REGION Network 189: CARRIER SPACING FAULT
   RUNG wire#powerrail
      Contact( "reset" )
      Contact( "EMS".Carrier[5].SDC_OUT.Faults.CarrierSpacingFault )
      wire#w1
      Coil( "DB302_HMI_Faults".Carrier5_Faults_2.%X2 )
   END_RUNG
   RUNG wire#powerrail
      Contact( "DB302_HMI_Faults".Carrier5_Faults_2.%X2 )
      I_Contact( "EMS_Fault_Reset" )
   END_RUNG wire#w1
   // the same network as SCL:
   "DB302_HMI_Faults".Carrier5_Faults_2.%X2 := ("reset" AND "EMS".Carrier[5].SDC_OUT.Faults.CarrierSpacingFault) OR ("DB302_HMI_Faults".Carrier5_Faults_2.%X2 AND NOT "EMS_Fault_Reset");
END_REGION

REGION Network 190: DUPLICATE CARRIER NUMBER FAULT
   RUNG wire#powerrail
      Contact( "reset" )
      Contact( "EMS".Carrier[5].SDC_OUT.Faults.DuplicateCarrierFault )
      wire#w1
      Coil( "DB302_HMI_Faults".Carrier5_Faults_2.%X3 )
   END_RUNG
   RUNG wire#powerrail
      Contact( "DB302_HMI_Faults".Carrier5_Faults_2.%X3 )
      I_Contact( "EMS_Fault_Reset" )
   END_RUNG wire#w1
   // the same network as SCL:
   "DB302_HMI_Faults".Carrier5_Faults_2.%X3 := ("reset" AND "EMS".Carrier[5].SDC_OUT.Faults.DuplicateCarrierFault) OR ("DB302_HMI_Faults".Carrier5_Faults_2.%X3 AND NOT "EMS_Fault_Reset");
END_REGION

REGION Network 191: PRODUCTION HOLD PB NOT RESET
   RUNG wire#powerrail
      Contact( "reset" )
      { S7_Templates := "SrcType := Word" } EQ_Contact(in1 := "DB101_DB_SDC_FAULTS".Carrier_Fault[5], in2 := 103)
      Coil( "DB302_HMI_Faults".Carrier5_Faults_3.%X14 )
   END_RUNG
   // the same network as SCL:
   "DB302_HMI_Faults".Carrier5_Faults_3.%X14 := "reset" AND ("DB101_DB_SDC_FAULTS".Carrier_Fault[5] = 103);
END_REGION

REGION Network 192: CARRIER FAULTS MASKED
   Label( C05_Comm_Flt )
   RUNG wire#powerrail
      Contact( "EMS".Carrier[5].FaultsMasked )
      Coil( "DB302_HMI_Faults".Carrier5_Faults_3.%X15 )
   END_RUNG
   // the same network as SCL:
   C05_Comm_Flt:
   "DB302_HMI_Faults".Carrier5_Faults_3.%X15 := "EMS".Carrier[5].FaultsMasked;
END_REGION

REGION Network 193: CARRIER 6 FAULTS
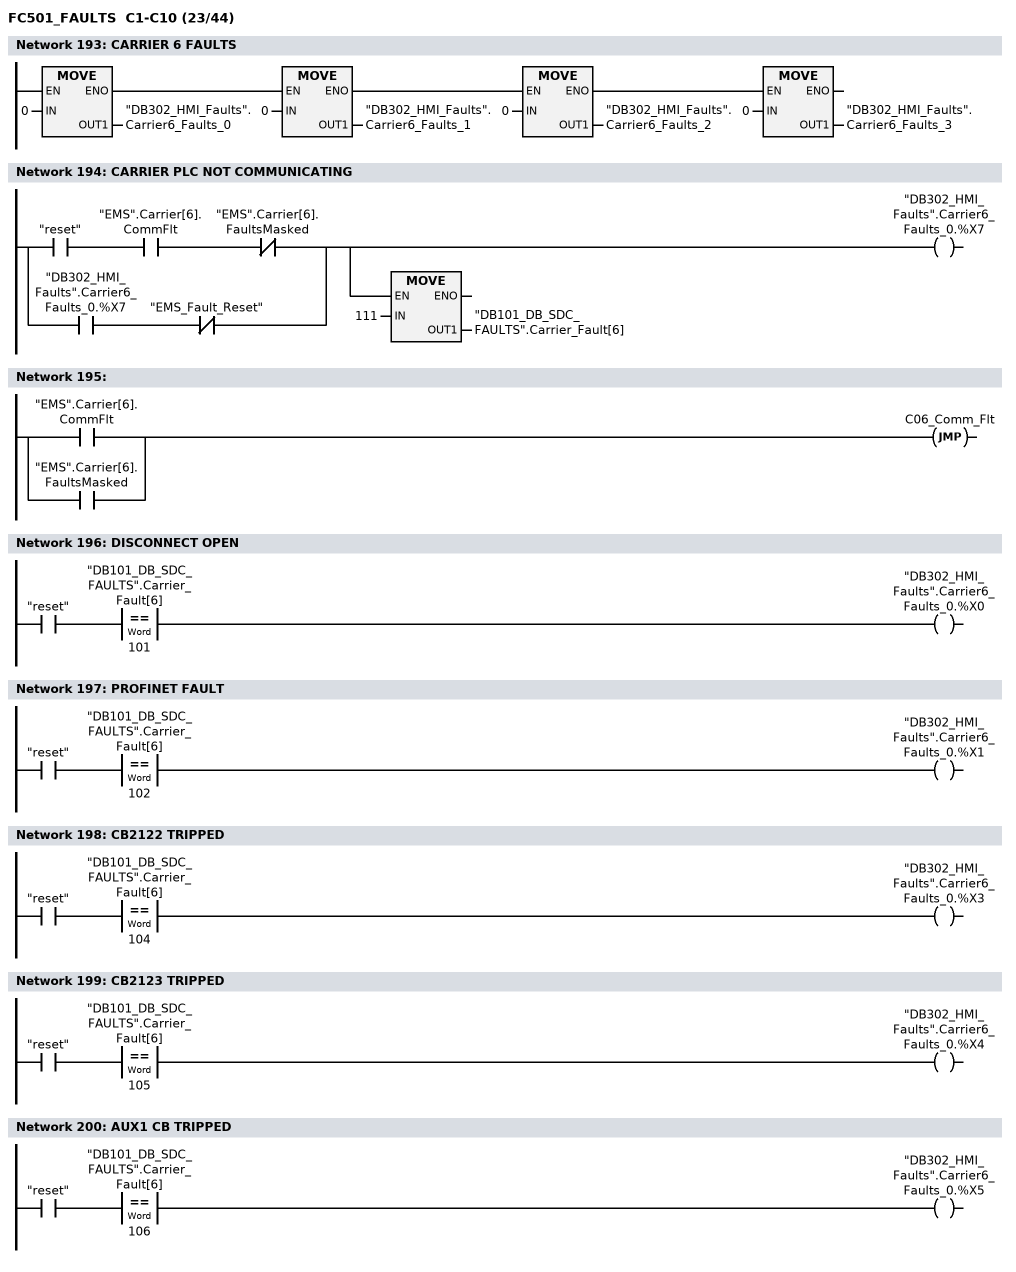
   RUNG wire#powerrail
      Move(in := 0, out1 => "DB302_HMI_Faults".Carrier6_Faults_0)
      Move(in := 0, out1 => "DB302_HMI_Faults".Carrier6_Faults_1)
      Move(in := 0, out1 => "DB302_HMI_Faults".Carrier6_Faults_2)
      Move(in := 0, out1 => "DB302_HMI_Faults".Carrier6_Faults_3)
   END_RUNG
   // the same network as SCL:
   "DB302_HMI_Faults".Carrier6_Faults_0 := 0;
   "DB302_HMI_Faults".Carrier6_Faults_1 := 0;
   "DB302_HMI_Faults".Carrier6_Faults_2 := 0;
   "DB302_HMI_Faults".Carrier6_Faults_3 := 0;
END_REGION

REGION Network 194: CARRIER PLC NOT COMMUNICATING
   RUNG wire#powerrail
      Contact( "reset" )
      Contact( "EMS".Carrier[6].CommFlt )
      I_Contact( "EMS".Carrier[6].FaultsMasked )
      wire#w1
      Coil( "DB302_HMI_Faults".Carrier6_Faults_0.%X7 )
   END_RUNG
   RUNG wire#powerrail
      Contact( "DB302_HMI_Faults".Carrier6_Faults_0.%X7 )
      I_Contact( "EMS_Fault_Reset" )
   END_RUNG wire#w1
   RUNG wire#w1
      Move(in := 111, out1 => "DB101_DB_SDC_FAULTS".Carrier_Fault[6])
   END_RUNG
   // the same network as SCL:
   "DB302_HMI_Faults".Carrier6_Faults_0.%X7 := ("reset" AND "EMS".Carrier[6].CommFlt AND NOT "EMS".Carrier[6].FaultsMasked) OR ("DB302_HMI_Faults".Carrier6_Faults_0.%X7 AND NOT "EMS_Fault_Reset");
   IF "DB302_HMI_Faults".Carrier6_Faults_0.%X7 THEN "DB101_DB_SDC_FAULTS".Carrier_Fault[6] := 111; END_IF;
END_REGION

REGION Network 195
   RUNG wire#powerrail
      Contact( "EMS".Carrier[6].CommFlt )
      wire#w1
      JumpCoil( C06_Comm_Flt )
   END_RUNG
   RUNG wire#powerrail
      Contact( "EMS".Carrier[6].FaultsMasked )
   END_RUNG wire#w1
   // the same network as SCL:
   IF "EMS".Carrier[6].CommFlt OR "EMS".Carrier[6].FaultsMasked THEN GOTO C06_Comm_Flt; END_IF;
END_REGION

REGION Network 196: DISCONNECT OPEN
   RUNG wire#powerrail
      Contact( "reset" )
      { S7_Templates := "SrcType := Word" } EQ_Contact(in1 := "DB101_DB_SDC_FAULTS".Carrier_Fault[6], in2 := 101)
      Coil( "DB302_HMI_Faults".Carrier6_Faults_0.%X0 )
   END_RUNG
   // the same network as SCL:
   "DB302_HMI_Faults".Carrier6_Faults_0.%X0 := "reset" AND ("DB101_DB_SDC_FAULTS".Carrier_Fault[6] = 101);
END_REGION

REGION Network 197: PROFINET FAULT
   RUNG wire#powerrail
      Contact( "reset" )
      { S7_Templates := "SrcType := Word" } EQ_Contact(in1 := "DB101_DB_SDC_FAULTS".Carrier_Fault[6], in2 := 102)
      Coil( "DB302_HMI_Faults".Carrier6_Faults_0.%X1 )
   END_RUNG
   // the same network as SCL:
   "DB302_HMI_Faults".Carrier6_Faults_0.%X1 := "reset" AND ("DB101_DB_SDC_FAULTS".Carrier_Fault[6] = 102);
END_REGION

REGION Network 198: CB2122 TRIPPED
   RUNG wire#powerrail
      Contact( "reset" )
      { S7_Templates := "SrcType := Word" } EQ_Contact(in1 := "DB101_DB_SDC_FAULTS".Carrier_Fault[6], in2 := 104)
      Coil( "DB302_HMI_Faults".Carrier6_Faults_0.%X3 )
   END_RUNG
   // the same network as SCL:
   "DB302_HMI_Faults".Carrier6_Faults_0.%X3 := "reset" AND ("DB101_DB_SDC_FAULTS".Carrier_Fault[6] = 104);
END_REGION

REGION Network 199: CB2123 TRIPPED
   RUNG wire#powerrail
      Contact( "reset" )
      { S7_Templates := "SrcType := Word" } EQ_Contact(in1 := "DB101_DB_SDC_FAULTS".Carrier_Fault[6], in2 := 105)
      Coil( "DB302_HMI_Faults".Carrier6_Faults_0.%X4 )
   END_RUNG
   // the same network as SCL:
   "DB302_HMI_Faults".Carrier6_Faults_0.%X4 := "reset" AND ("DB101_DB_SDC_FAULTS".Carrier_Fault[6] = 105);
END_REGION

REGION Network 200: AUX1 CB TRIPPED
   RUNG wire#powerrail
      Contact( "reset" )
      { S7_Templates := "SrcType := Word" } EQ_Contact(in1 := "DB101_DB_SDC_FAULTS".Carrier_Fault[6], in2 := 106)
      Coil( "DB302_HMI_Faults".Carrier6_Faults_0.%X5 )
   END_RUNG
   // the same network as SCL:
   "DB302_HMI_Faults".Carrier6_Faults_0.%X5 := "reset" AND ("DB101_DB_SDC_FAULTS".Carrier_Fault[6] = 106);
END_REGION

REGION Network 201: AUX2 CB TRIPPED
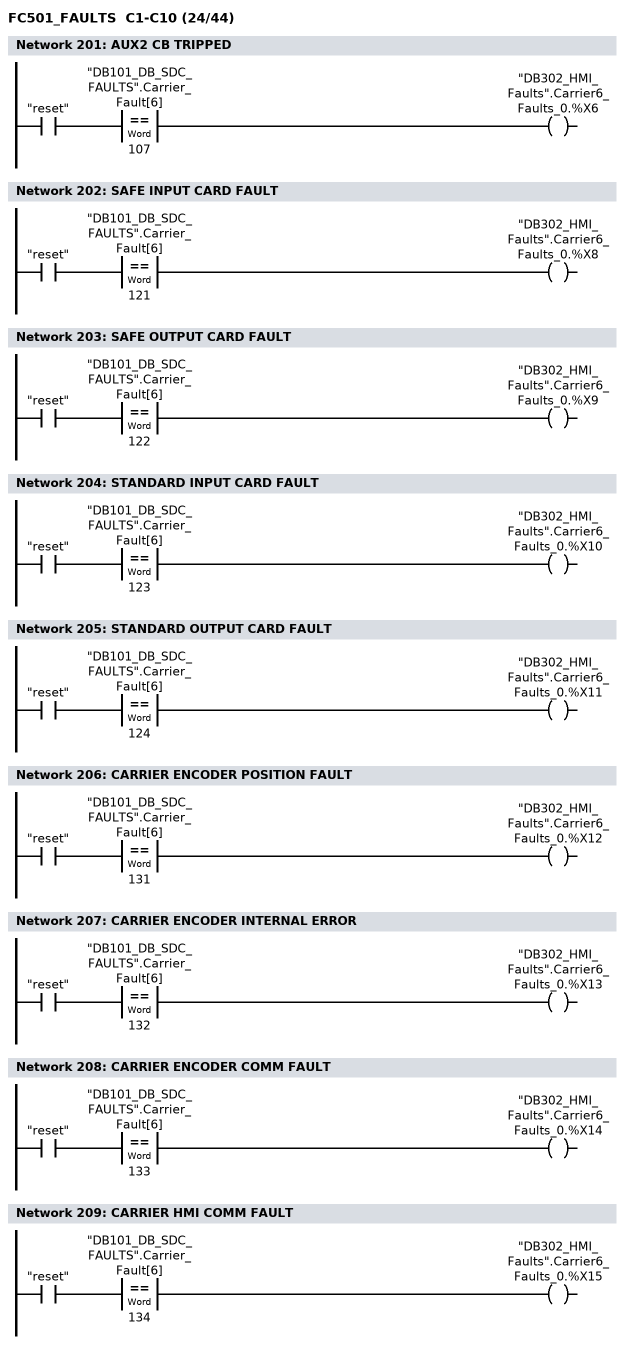
   RUNG wire#powerrail
      Contact( "reset" )
      { S7_Templates := "SrcType := Word" } EQ_Contact(in1 := "DB101_DB_SDC_FAULTS".Carrier_Fault[6], in2 := 107)
      Coil( "DB302_HMI_Faults".Carrier6_Faults_0.%X6 )
   END_RUNG
   // the same network as SCL:
   "DB302_HMI_Faults".Carrier6_Faults_0.%X6 := "reset" AND ("DB101_DB_SDC_FAULTS".Carrier_Fault[6] = 107);
END_REGION

REGION Network 202: SAFE INPUT CARD FAULT
   RUNG wire#powerrail
      Contact( "reset" )
      { S7_Templates := "SrcType := Word" } EQ_Contact(in1 := "DB101_DB_SDC_FAULTS".Carrier_Fault[6], in2 := 121)
      Coil( "DB302_HMI_Faults".Carrier6_Faults_0.%X8 )
   END_RUNG
   // the same network as SCL:
   "DB302_HMI_Faults".Carrier6_Faults_0.%X8 := "reset" AND ("DB101_DB_SDC_FAULTS".Carrier_Fault[6] = 121);
END_REGION

REGION Network 203: SAFE OUTPUT CARD FAULT
   RUNG wire#powerrail
      Contact( "reset" )
      { S7_Templates := "SrcType := Word" } EQ_Contact(in1 := "DB101_DB_SDC_FAULTS".Carrier_Fault[6], in2 := 122)
      Coil( "DB302_HMI_Faults".Carrier6_Faults_0.%X9 )
   END_RUNG
   // the same network as SCL:
   "DB302_HMI_Faults".Carrier6_Faults_0.%X9 := "reset" AND ("DB101_DB_SDC_FAULTS".Carrier_Fault[6] = 122);
END_REGION

REGION Network 204: STANDARD INPUT CARD FAULT
   RUNG wire#powerrail
      Contact( "reset" )
      { S7_Templates := "SrcType := Word" } EQ_Contact(in1 := "DB101_DB_SDC_FAULTS".Carrier_Fault[6], in2 := 123)
      Coil( "DB302_HMI_Faults".Carrier6_Faults_0.%X10 )
   END_RUNG
   // the same network as SCL:
   "DB302_HMI_Faults".Carrier6_Faults_0.%X10 := "reset" AND ("DB101_DB_SDC_FAULTS".Carrier_Fault[6] = 123);
END_REGION

REGION Network 205: STANDARD OUTPUT CARD FAULT
   RUNG wire#powerrail
      Contact( "reset" )
      { S7_Templates := "SrcType := Word" } EQ_Contact(in1 := "DB101_DB_SDC_FAULTS".Carrier_Fault[6], in2 := 124)
      Coil( "DB302_HMI_Faults".Carrier6_Faults_0.%X11 )
   END_RUNG
   // the same network as SCL:
   "DB302_HMI_Faults".Carrier6_Faults_0.%X11 := "reset" AND ("DB101_DB_SDC_FAULTS".Carrier_Fault[6] = 124);
END_REGION

REGION Network 206: CARRIER ENCODER POSITION FAULT
   RUNG wire#powerrail
      Contact( "reset" )
      { S7_Templates := "SrcType := Word" } EQ_Contact(in1 := "DB101_DB_SDC_FAULTS".Carrier_Fault[6], in2 := 131)
      Coil( "DB302_HMI_Faults".Carrier6_Faults_0.%X12 )
   END_RUNG
   // the same network as SCL:
   "DB302_HMI_Faults".Carrier6_Faults_0.%X12 := "reset" AND ("DB101_DB_SDC_FAULTS".Carrier_Fault[6] = 131);
END_REGION

REGION Network 207: CARRIER ENCODER INTERNAL ERROR
   RUNG wire#powerrail
      Contact( "reset" )
      { S7_Templates := "SrcType := Word" } EQ_Contact(in1 := "DB101_DB_SDC_FAULTS".Carrier_Fault[6], in2 := 132)
      Coil( "DB302_HMI_Faults".Carrier6_Faults_0.%X13 )
   END_RUNG
   // the same network as SCL:
   "DB302_HMI_Faults".Carrier6_Faults_0.%X13 := "reset" AND ("DB101_DB_SDC_FAULTS".Carrier_Fault[6] = 132);
END_REGION

REGION Network 208: CARRIER ENCODER COMM FAULT
   RUNG wire#powerrail
      Contact( "reset" )
      { S7_Templates := "SrcType := Word" } EQ_Contact(in1 := "DB101_DB_SDC_FAULTS".Carrier_Fault[6], in2 := 133)
      Coil( "DB302_HMI_Faults".Carrier6_Faults_0.%X14 )
   END_RUNG
   // the same network as SCL:
   "DB302_HMI_Faults".Carrier6_Faults_0.%X14 := "reset" AND ("DB101_DB_SDC_FAULTS".Carrier_Fault[6] = 133);
END_REGION

REGION Network 209: CARRIER HMI COMM FAULT
   RUNG wire#powerrail
      Contact( "reset" )
      { S7_Templates := "SrcType := Word" } EQ_Contact(in1 := "DB101_DB_SDC_FAULTS".Carrier_Fault[6], in2 := 134)
      Coil( "DB302_HMI_Faults".Carrier6_Faults_0.%X15 )
   END_RUNG
   // the same network as SCL:
   "DB302_HMI_Faults".Carrier6_Faults_0.%X15 := "reset" AND ("DB101_DB_SDC_FAULTS".Carrier_Fault[6] = 134);
END_REGION

REGION Network 210: CARRIER CRASH DETECTION FAULT
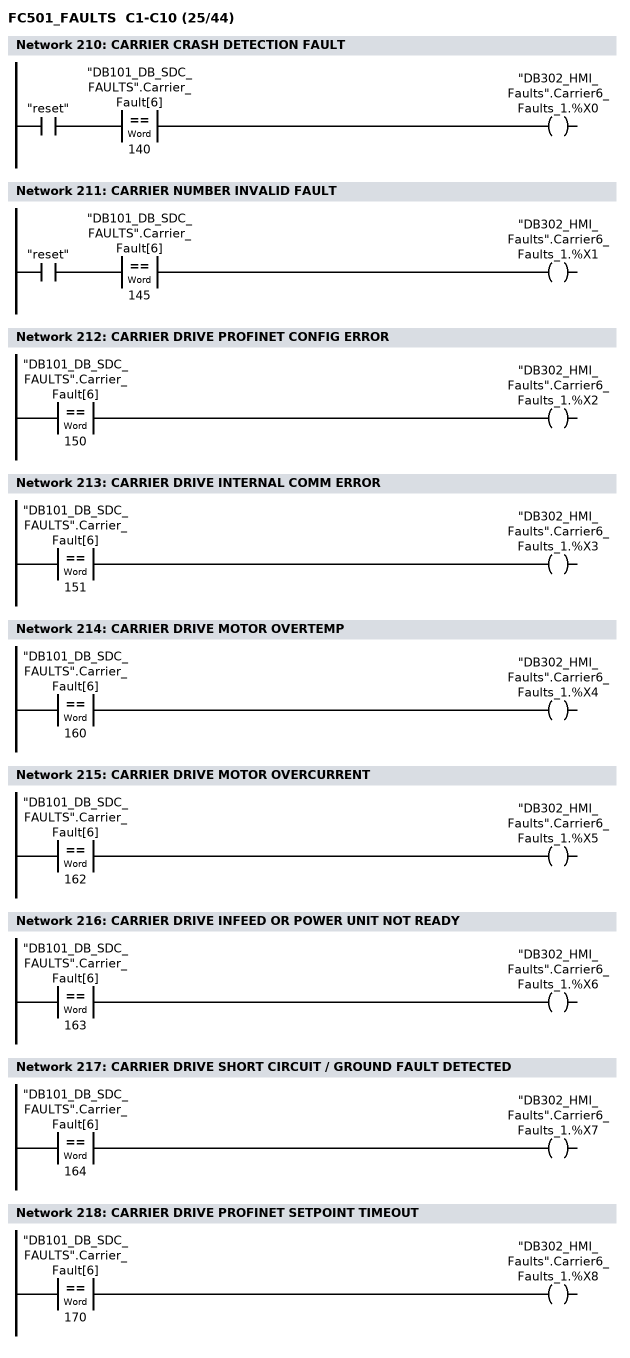
   RUNG wire#powerrail
      Contact( "reset" )
      { S7_Templates := "SrcType := Word" } EQ_Contact(in1 := "DB101_DB_SDC_FAULTS".Carrier_Fault[6], in2 := 140)
      Coil( "DB302_HMI_Faults".Carrier6_Faults_1.%X0 )
   END_RUNG
   // the same network as SCL:
   "DB302_HMI_Faults".Carrier6_Faults_1.%X0 := "reset" AND ("DB101_DB_SDC_FAULTS".Carrier_Fault[6] = 140);
END_REGION

REGION Network 211: CARRIER NUMBER INVALID FAULT
   RUNG wire#powerrail
      Contact( "reset" )
      { S7_Templates := "SrcType := Word" } EQ_Contact(in1 := "DB101_DB_SDC_FAULTS".Carrier_Fault[6], in2 := 145)
      Coil( "DB302_HMI_Faults".Carrier6_Faults_1.%X1 )
   END_RUNG
   // the same network as SCL:
   "DB302_HMI_Faults".Carrier6_Faults_1.%X1 := "reset" AND ("DB101_DB_SDC_FAULTS".Carrier_Fault[6] = 145);
END_REGION

REGION Network 212: CARRIER DRIVE PROFINET CONFIG ERROR
   RUNG wire#powerrail
      { S7_Templates := "SrcType := Word" } EQ_Contact(in1 := "DB101_DB_SDC_FAULTS".Carrier_Fault[6], in2 := 150)
      Coil( "DB302_HMI_Faults".Carrier6_Faults_1.%X2 )
   END_RUNG
   // the same network as SCL:
   "DB302_HMI_Faults".Carrier6_Faults_1.%X2 := "DB101_DB_SDC_FAULTS".Carrier_Fault[6] = 150;
END_REGION

REGION Network 213: CARRIER DRIVE INTERNAL COMM ERROR
   RUNG wire#powerrail
      { S7_Templates := "SrcType := Word" } EQ_Contact(in1 := "DB101_DB_SDC_FAULTS".Carrier_Fault[6], in2 := 151)
      Coil( "DB302_HMI_Faults".Carrier6_Faults_1.%X3 )
   END_RUNG
   // the same network as SCL:
   "DB302_HMI_Faults".Carrier6_Faults_1.%X3 := "DB101_DB_SDC_FAULTS".Carrier_Fault[6] = 151;
END_REGION

REGION Network 214: CARRIER DRIVE MOTOR OVERTEMP
   RUNG wire#powerrail
      { S7_Templates := "SrcType := Word" } EQ_Contact(in1 := "DB101_DB_SDC_FAULTS".Carrier_Fault[6], in2 := 160)
      Coil( "DB302_HMI_Faults".Carrier6_Faults_1.%X4 )
   END_RUNG
   // the same network as SCL:
   "DB302_HMI_Faults".Carrier6_Faults_1.%X4 := "DB101_DB_SDC_FAULTS".Carrier_Fault[6] = 160;
END_REGION

REGION Network 215: CARRIER DRIVE MOTOR OVERCURRENT
   RUNG wire#powerrail
      { S7_Templates := "SrcType := Word" } EQ_Contact(in1 := "DB101_DB_SDC_FAULTS".Carrier_Fault[6], in2 := 162)
      Coil( "DB302_HMI_Faults".Carrier6_Faults_1.%X5 )
   END_RUNG
   // the same network as SCL:
   "DB302_HMI_Faults".Carrier6_Faults_1.%X5 := "DB101_DB_SDC_FAULTS".Carrier_Fault[6] = 162;
END_REGION

REGION Network 216: CARRIER DRIVE INFEED OR POWER UNIT NOT READY
   RUNG wire#powerrail
      { S7_Templates := "SrcType := Word" } EQ_Contact(in1 := "DB101_DB_SDC_FAULTS".Carrier_Fault[6], in2 := 163)
      Coil( "DB302_HMI_Faults".Carrier6_Faults_1.%X6 )
   END_RUNG
   // the same network as SCL:
   "DB302_HMI_Faults".Carrier6_Faults_1.%X6 := "DB101_DB_SDC_FAULTS".Carrier_Fault[6] = 163;
END_REGION

REGION Network 217: CARRIER DRIVE SHORT CIRCUIT / GROUND FAULT DETECTED
   RUNG wire#powerrail
      { S7_Templates := "SrcType := Word" } EQ_Contact(in1 := "DB101_DB_SDC_FAULTS".Carrier_Fault[6], in2 := 164)
      Coil( "DB302_HMI_Faults".Carrier6_Faults_1.%X7 )
   END_RUNG
   // the same network as SCL:
   "DB302_HMI_Faults".Carrier6_Faults_1.%X7 := "DB101_DB_SDC_FAULTS".Carrier_Fault[6] = 164;
END_REGION

REGION Network 218: CARRIER DRIVE PROFINET SETPOINT TIMEOUT
   RUNG wire#powerrail
      { S7_Templates := "SrcType := Word" } EQ_Contact(in1 := "DB101_DB_SDC_FAULTS".Carrier_Fault[6], in2 := 170)
      Coil( "DB302_HMI_Faults".Carrier6_Faults_1.%X8 )
   END_RUNG
   // the same network as SCL:
   "DB302_HMI_Faults".Carrier6_Faults_1.%X8 := "DB101_DB_SDC_FAULTS".Carrier_Fault[6] = 170;
END_REGION

REGION Network 219: CARRIER POWER UNIT OVERCURRENT
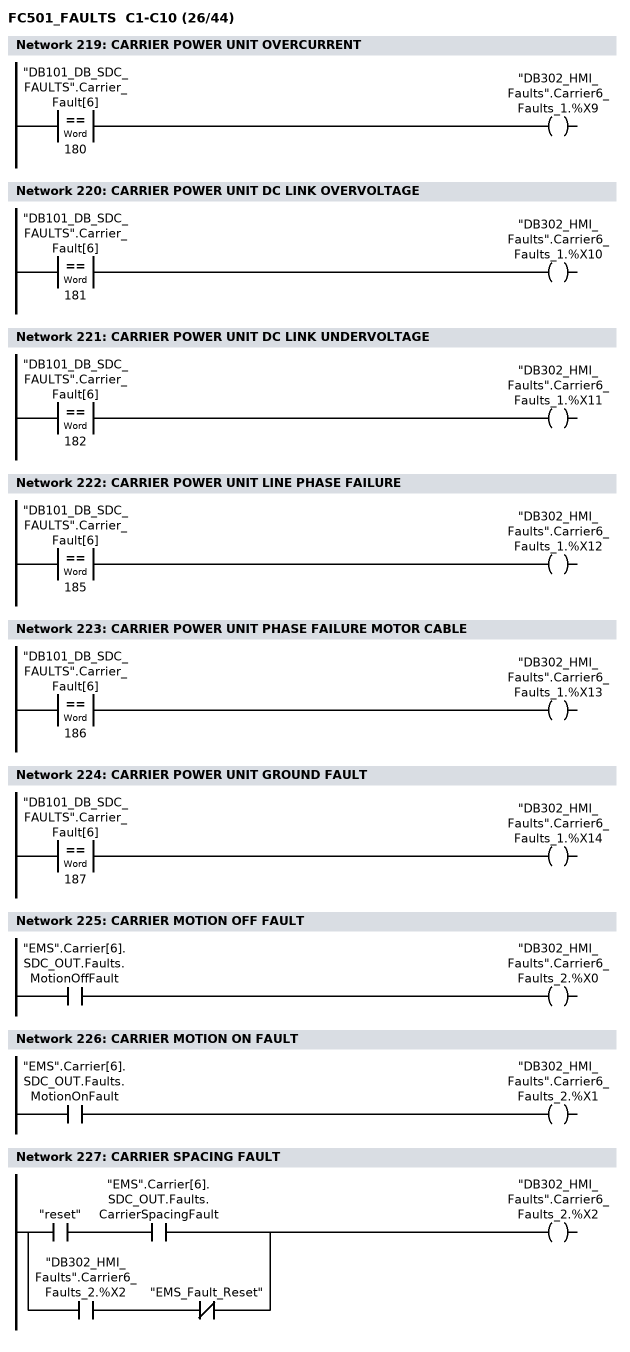
   RUNG wire#powerrail
      { S7_Templates := "SrcType := Word" } EQ_Contact(in1 := "DB101_DB_SDC_FAULTS".Carrier_Fault[6], in2 := 180)
      Coil( "DB302_HMI_Faults".Carrier6_Faults_1.%X9 )
   END_RUNG
   // the same network as SCL:
   "DB302_HMI_Faults".Carrier6_Faults_1.%X9 := "DB101_DB_SDC_FAULTS".Carrier_Fault[6] = 180;
END_REGION

REGION Network 220: CARRIER POWER UNIT DC LINK OVERVOLTAGE
   RUNG wire#powerrail
      { S7_Templates := "SrcType := Word" } EQ_Contact(in1 := "DB101_DB_SDC_FAULTS".Carrier_Fault[6], in2 := 181)
      Coil( "DB302_HMI_Faults".Carrier6_Faults_1.%X10 )
   END_RUNG
   // the same network as SCL:
   "DB302_HMI_Faults".Carrier6_Faults_1.%X10 := "DB101_DB_SDC_FAULTS".Carrier_Fault[6] = 181;
END_REGION

REGION Network 221: CARRIER POWER UNIT DC LINK UNDERVOLTAGE
   RUNG wire#powerrail
      { S7_Templates := "SrcType := Word" } EQ_Contact(in1 := "DB101_DB_SDC_FAULTS".Carrier_Fault[6], in2 := 182)
      Coil( "DB302_HMI_Faults".Carrier6_Faults_1.%X11 )
   END_RUNG
   // the same network as SCL:
   "DB302_HMI_Faults".Carrier6_Faults_1.%X11 := "DB101_DB_SDC_FAULTS".Carrier_Fault[6] = 182;
END_REGION

REGION Network 222: CARRIER POWER UNIT LINE PHASE FAILURE
   RUNG wire#powerrail
      { S7_Templates := "SrcType := Word" } EQ_Contact(in1 := "DB101_DB_SDC_FAULTS".Carrier_Fault[6], in2 := 185)
      Coil( "DB302_HMI_Faults".Carrier6_Faults_1.%X12 )
   END_RUNG
   // the same network as SCL:
   "DB302_HMI_Faults".Carrier6_Faults_1.%X12 := "DB101_DB_SDC_FAULTS".Carrier_Fault[6] = 185;
END_REGION

REGION Network 223: CARRIER POWER UNIT PHASE FAILURE MOTOR CABLE
   RUNG wire#powerrail
      { S7_Templates := "SrcType := Word" } EQ_Contact(in1 := "DB101_DB_SDC_FAULTS".Carrier_Fault[6], in2 := 186)
      Coil( "DB302_HMI_Faults".Carrier6_Faults_1.%X13 )
   END_RUNG
   // the same network as SCL:
   "DB302_HMI_Faults".Carrier6_Faults_1.%X13 := "DB101_DB_SDC_FAULTS".Carrier_Fault[6] = 186;
END_REGION

REGION Network 224: CARRIER POWER UNIT GROUND FAULT
   RUNG wire#powerrail
      { S7_Templates := "SrcType := Word" } EQ_Contact(in1 := "DB101_DB_SDC_FAULTS".Carrier_Fault[6], in2 := 187)
      Coil( "DB302_HMI_Faults".Carrier6_Faults_1.%X14 )
   END_RUNG
   // the same network as SCL:
   "DB302_HMI_Faults".Carrier6_Faults_1.%X14 := "DB101_DB_SDC_FAULTS".Carrier_Fault[6] = 187;
END_REGION

REGION Network 225: CARRIER MOTION OFF FAULT
   RUNG wire#powerrail
      Contact( "EMS".Carrier[6].SDC_OUT.Faults.MotionOffFault )
      Coil( "DB302_HMI_Faults".Carrier6_Faults_2.%X0 )
   END_RUNG
   // the same network as SCL:
   "DB302_HMI_Faults".Carrier6_Faults_2.%X0 := "EMS".Carrier[6].SDC_OUT.Faults.MotionOffFault;
END_REGION

REGION Network 226: CARRIER MOTION ON FAULT
   RUNG wire#powerrail
      Contact( "EMS".Carrier[6].SDC_OUT.Faults.MotionOnFault )
      Coil( "DB302_HMI_Faults".Carrier6_Faults_2.%X1 )
   END_RUNG
   // the same network as SCL:
   "DB302_HMI_Faults".Carrier6_Faults_2.%X1 := "EMS".Carrier[6].SDC_OUT.Faults.MotionOnFault;
END_REGION

REGION Network 227: CARRIER SPACING FAULT
   RUNG wire#powerrail
      Contact( "reset" )
      Contact( "EMS".Carrier[6].SDC_OUT.Faults.CarrierSpacingFault )
      wire#w1
      Coil( "DB302_HMI_Faults".Carrier6_Faults_2.%X2 )
   END_RUNG
   RUNG wire#powerrail
      Contact( "DB302_HMI_Faults".Carrier6_Faults_2.%X2 )
      I_Contact( "EMS_Fault_Reset" )
   END_RUNG wire#w1
   // the same network as SCL:
   "DB302_HMI_Faults".Carrier6_Faults_2.%X2 := ("reset" AND "EMS".Carrier[6].SDC_OUT.Faults.CarrierSpacingFault) OR ("DB302_HMI_Faults".Carrier6_Faults_2.%X2 AND NOT "EMS_Fault_Reset");
END_REGION

REGION Network 228: DUPLICATE CARRIER NUMBER FAULT
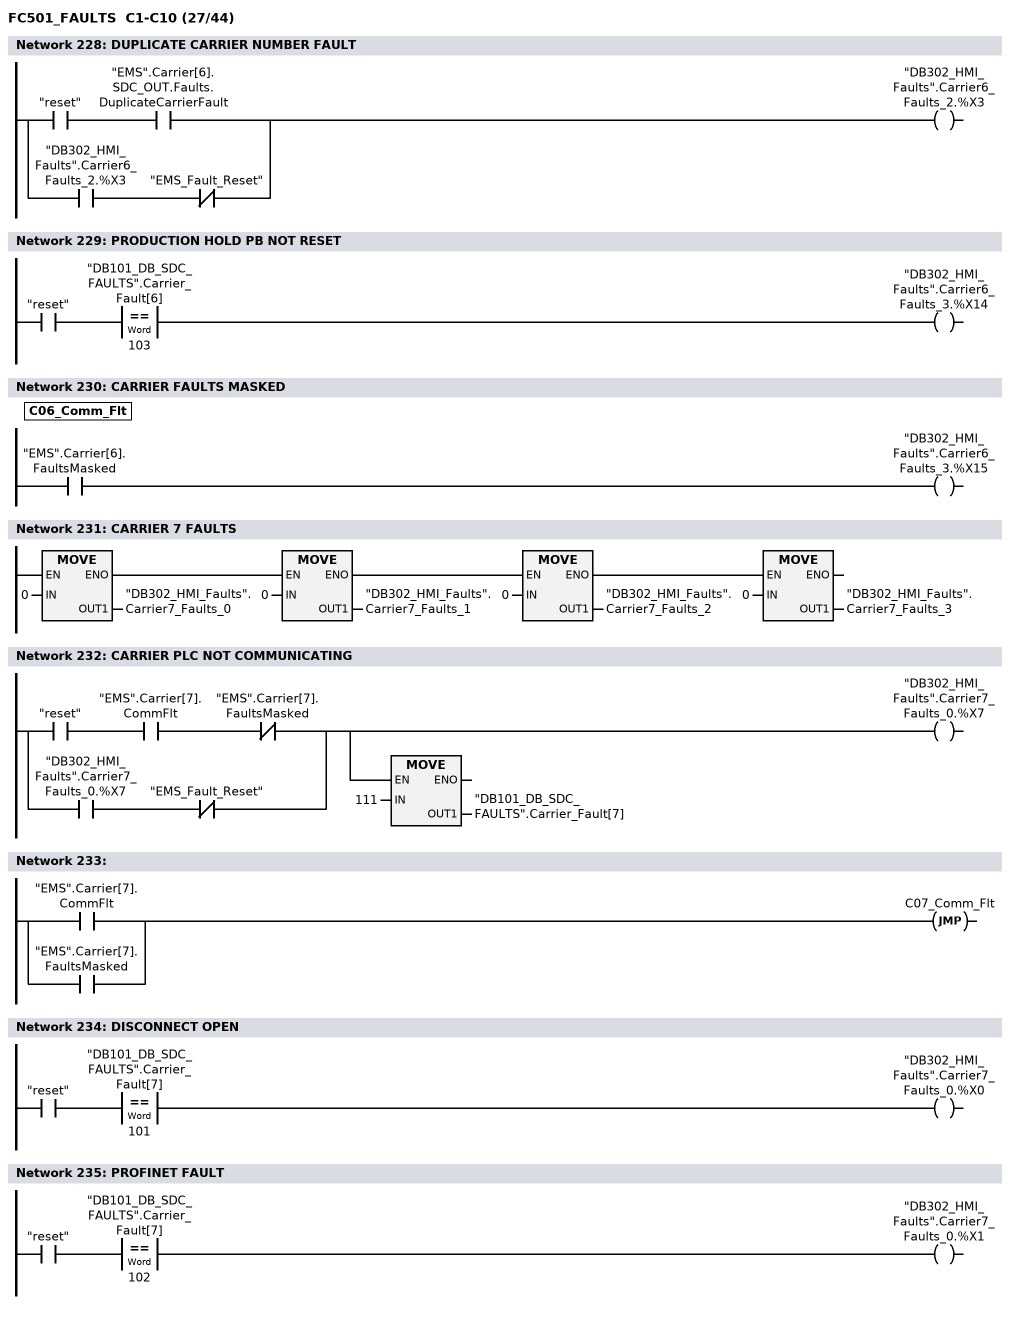
   RUNG wire#powerrail
      Contact( "reset" )
      Contact( "EMS".Carrier[6].SDC_OUT.Faults.DuplicateCarrierFault )
      wire#w1
      Coil( "DB302_HMI_Faults".Carrier6_Faults_2.%X3 )
   END_RUNG
   RUNG wire#powerrail
      Contact( "DB302_HMI_Faults".Carrier6_Faults_2.%X3 )
      I_Contact( "EMS_Fault_Reset" )
   END_RUNG wire#w1
   // the same network as SCL:
   "DB302_HMI_Faults".Carrier6_Faults_2.%X3 := ("reset" AND "EMS".Carrier[6].SDC_OUT.Faults.DuplicateCarrierFault) OR ("DB302_HMI_Faults".Carrier6_Faults_2.%X3 AND NOT "EMS_Fault_Reset");
END_REGION

REGION Network 229: PRODUCTION HOLD PB NOT RESET
   RUNG wire#powerrail
      Contact( "reset" )
      { S7_Templates := "SrcType := Word" } EQ_Contact(in1 := "DB101_DB_SDC_FAULTS".Carrier_Fault[6], in2 := 103)
      Coil( "DB302_HMI_Faults".Carrier6_Faults_3.%X14 )
   END_RUNG
   // the same network as SCL:
   "DB302_HMI_Faults".Carrier6_Faults_3.%X14 := "reset" AND ("DB101_DB_SDC_FAULTS".Carrier_Fault[6] = 103);
END_REGION

REGION Network 230: CARRIER FAULTS MASKED
   Label( C06_Comm_Flt )
   RUNG wire#powerrail
      Contact( "EMS".Carrier[6].FaultsMasked )
      Coil( "DB302_HMI_Faults".Carrier6_Faults_3.%X15 )
   END_RUNG
   // the same network as SCL:
   C06_Comm_Flt:
   "DB302_HMI_Faults".Carrier6_Faults_3.%X15 := "EMS".Carrier[6].FaultsMasked;
END_REGION

REGION Network 231: CARRIER 7 FAULTS
   RUNG wire#powerrail
      Move(in := 0, out1 => "DB302_HMI_Faults".Carrier7_Faults_0)
      Move(in := 0, out1 => "DB302_HMI_Faults".Carrier7_Faults_1)
      Move(in := 0, out1 => "DB302_HMI_Faults".Carrier7_Faults_2)
      Move(in := 0, out1 => "DB302_HMI_Faults".Carrier7_Faults_3)
   END_RUNG
   // the same network as SCL:
   "DB302_HMI_Faults".Carrier7_Faults_0 := 0;
   "DB302_HMI_Faults".Carrier7_Faults_1 := 0;
   "DB302_HMI_Faults".Carrier7_Faults_2 := 0;
   "DB302_HMI_Faults".Carrier7_Faults_3 := 0;
END_REGION

REGION Network 232: CARRIER PLC NOT COMMUNICATING
   RUNG wire#powerrail
      Contact( "reset" )
      Contact( "EMS".Carrier[7].CommFlt )
      I_Contact( "EMS".Carrier[7].FaultsMasked )
      wire#w1
      Coil( "DB302_HMI_Faults".Carrier7_Faults_0.%X7 )
   END_RUNG
   RUNG wire#powerrail
      Contact( "DB302_HMI_Faults".Carrier7_Faults_0.%X7 )
      I_Contact( "EMS_Fault_Reset" )
   END_RUNG wire#w1
   RUNG wire#w1
      Move(in := 111, out1 => "DB101_DB_SDC_FAULTS".Carrier_Fault[7])
   END_RUNG
   // the same network as SCL:
   "DB302_HMI_Faults".Carrier7_Faults_0.%X7 := ("reset" AND "EMS".Carrier[7].CommFlt AND NOT "EMS".Carrier[7].FaultsMasked) OR ("DB302_HMI_Faults".Carrier7_Faults_0.%X7 AND NOT "EMS_Fault_Reset");
   IF "DB302_HMI_Faults".Carrier7_Faults_0.%X7 THEN "DB101_DB_SDC_FAULTS".Carrier_Fault[7] := 111; END_IF;
END_REGION

REGION Network 233
   RUNG wire#powerrail
      Contact( "EMS".Carrier[7].CommFlt )
      wire#w1
      JumpCoil( C07_Comm_Flt )
   END_RUNG
   RUNG wire#powerrail
      Contact( "EMS".Carrier[7].FaultsMasked )
   END_RUNG wire#w1
   // the same network as SCL:
   IF "EMS".Carrier[7].CommFlt OR "EMS".Carrier[7].FaultsMasked THEN GOTO C07_Comm_Flt; END_IF;
END_REGION

REGION Network 234: DISCONNECT OPEN
   RUNG wire#powerrail
      Contact( "reset" )
      { S7_Templates := "SrcType := Word" } EQ_Contact(in1 := "DB101_DB_SDC_FAULTS".Carrier_Fault[7], in2 := 101)
      Coil( "DB302_HMI_Faults".Carrier7_Faults_0.%X0 )
   END_RUNG
   // the same network as SCL:
   "DB302_HMI_Faults".Carrier7_Faults_0.%X0 := "reset" AND ("DB101_DB_SDC_FAULTS".Carrier_Fault[7] = 101);
END_REGION

REGION Network 235: PROFINET FAULT
   RUNG wire#powerrail
      Contact( "reset" )
      { S7_Templates := "SrcType := Word" } EQ_Contact(in1 := "DB101_DB_SDC_FAULTS".Carrier_Fault[7], in2 := 102)
      Coil( "DB302_HMI_Faults".Carrier7_Faults_0.%X1 )
   END_RUNG
   // the same network as SCL:
   "DB302_HMI_Faults".Carrier7_Faults_0.%X1 := "reset" AND ("DB101_DB_SDC_FAULTS".Carrier_Fault[7] = 102);
END_REGION

REGION Network 236: CB2122 TRIPPED
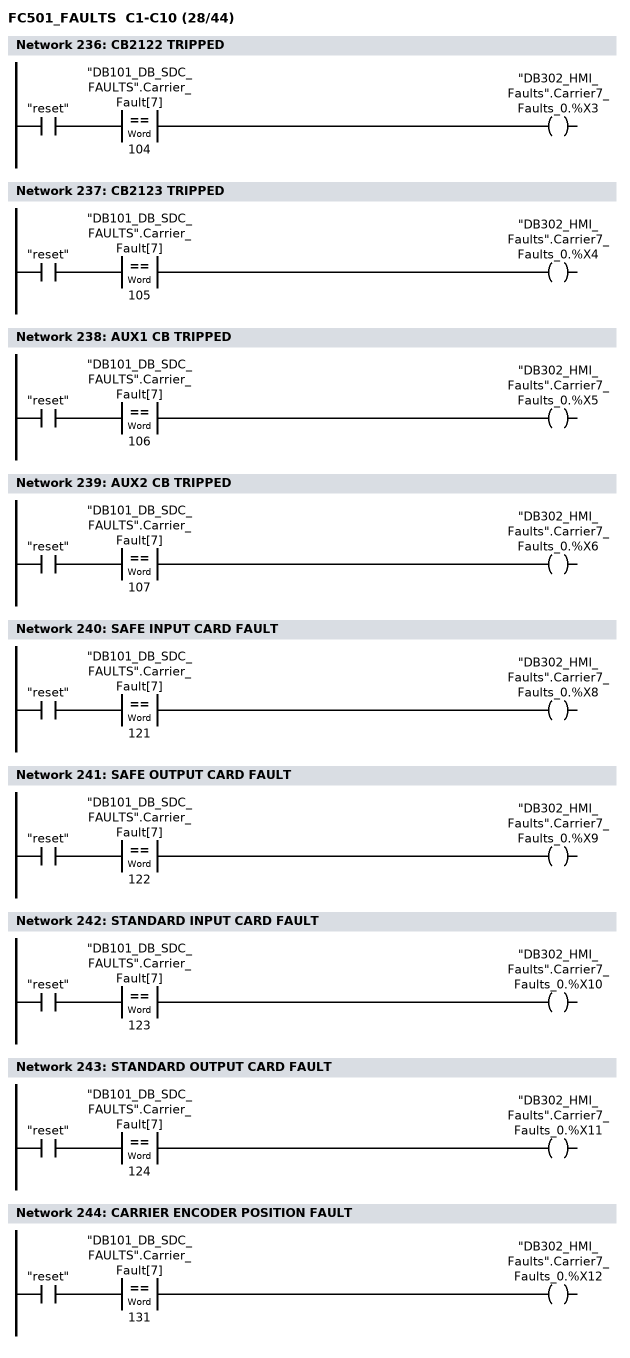
   RUNG wire#powerrail
      Contact( "reset" )
      { S7_Templates := "SrcType := Word" } EQ_Contact(in1 := "DB101_DB_SDC_FAULTS".Carrier_Fault[7], in2 := 104)
      Coil( "DB302_HMI_Faults".Carrier7_Faults_0.%X3 )
   END_RUNG
   // the same network as SCL:
   "DB302_HMI_Faults".Carrier7_Faults_0.%X3 := "reset" AND ("DB101_DB_SDC_FAULTS".Carrier_Fault[7] = 104);
END_REGION

REGION Network 237: CB2123 TRIPPED
   RUNG wire#powerrail
      Contact( "reset" )
      { S7_Templates := "SrcType := Word" } EQ_Contact(in1 := "DB101_DB_SDC_FAULTS".Carrier_Fault[7], in2 := 105)
      Coil( "DB302_HMI_Faults".Carrier7_Faults_0.%X4 )
   END_RUNG
   // the same network as SCL:
   "DB302_HMI_Faults".Carrier7_Faults_0.%X4 := "reset" AND ("DB101_DB_SDC_FAULTS".Carrier_Fault[7] = 105);
END_REGION

REGION Network 238: AUX1 CB TRIPPED
   RUNG wire#powerrail
      Contact( "reset" )
      { S7_Templates := "SrcType := Word" } EQ_Contact(in1 := "DB101_DB_SDC_FAULTS".Carrier_Fault[7], in2 := 106)
      Coil( "DB302_HMI_Faults".Carrier7_Faults_0.%X5 )
   END_RUNG
   // the same network as SCL:
   "DB302_HMI_Faults".Carrier7_Faults_0.%X5 := "reset" AND ("DB101_DB_SDC_FAULTS".Carrier_Fault[7] = 106);
END_REGION

REGION Network 239: AUX2 CB TRIPPED
   RUNG wire#powerrail
      Contact( "reset" )
      { S7_Templates := "SrcType := Word" } EQ_Contact(in1 := "DB101_DB_SDC_FAULTS".Carrier_Fault[7], in2 := 107)
      Coil( "DB302_HMI_Faults".Carrier7_Faults_0.%X6 )
   END_RUNG
   // the same network as SCL:
   "DB302_HMI_Faults".Carrier7_Faults_0.%X6 := "reset" AND ("DB101_DB_SDC_FAULTS".Carrier_Fault[7] = 107);
END_REGION

REGION Network 240: SAFE INPUT CARD FAULT
   RUNG wire#powerrail
      Contact( "reset" )
      { S7_Templates := "SrcType := Word" } EQ_Contact(in1 := "DB101_DB_SDC_FAULTS".Carrier_Fault[7], in2 := 121)
      Coil( "DB302_HMI_Faults".Carrier7_Faults_0.%X8 )
   END_RUNG
   // the same network as SCL:
   "DB302_HMI_Faults".Carrier7_Faults_0.%X8 := "reset" AND ("DB101_DB_SDC_FAULTS".Carrier_Fault[7] = 121);
END_REGION
